VERSION : 0.1
   STRUCT
      CarrierNumber : Word;
      CarrierPosition : DWord;
      ActualSpeed : Word;
      CarrierDriveFaults : Word;
      CarrierDriveAlarms : Word;
      CarrierFaults : Word;
      Spare_Word : Word;
      RunningFWD : Bool;
      RunningREV : Bool;
      Stopped : Bool;
      ProductionHoldPB_Status : Bool;
      CrashDetectStatus : Bool;
      HeartBeat : Bool;
      AutoMode : Bool;
      ManualMode : Bool;
      IR_Remote_9_Pressed : Bool;
      EncoderCommFault : Bool;
      DriveCommFault : Bool;
      HMICommFault : Bool;
   END_STRUCT;
END_TYPE

TYPE "UDT_SDC_OUT"
VERSION : 0.1
   STRUCT
      Zone : Int;
      CarrierNum : Word;
      CarrierPosition : DWord;
      NextCarrierNum : Word;
      NextStopPos : DWord;
      DriveFwdCMD : Bool;
      DriveCmdSpeed : Word;
      Spare_Word_1 : Word;
      Spare_Word_2 : Word;
      HeartBeat : Bool;
      FaultReset : Bool;
      HighSpeedEnable : Bool;
      AtCmdPos : Bool;
      DuplicateCarrierNum : Word;
      FirstDuplicateFndPos : Bool;
      SecondDuplicateFndPos : Bool;
      Faults : "UDT_SDCOutFaults";
   END_STRUCT;
END_TYPE

TYPE "UDT_CarrierFaults"
VERSION : 0.1
   STRUCT
      Fault : Array[0..9] of Int;
   END_STRUCT;
END_TYPE

TYPE "UDT_SDC"
   STRUCT
      HMI : "UDT_Drive_HMI";
   END_STRUCT;
END_TYPE

TYPE "UDT_TrafficCop"
VERSION : 0.1
   STRUCT
      Element_1 : Bool;
      AutoSpeedFast : Word;
      AutoSpeedSlow : Word;
      CommandPosLowLimit : DWord;
      CommandPosHighLimit : DWord;
      CommandPos : DWord;
      AtCommandPos : Bool;
      DecelPosition : DWord;
   END_STRUCT;
END_TYPE

TYPE "UDT_SDC_6EMS_TS_STAT"
VERSION : 0.1
   STRUCT
      EMS : Array[1..6] of "UDT_SDC_EMS_TS_STAT";
   END_STRUCT;
END_TYPE

TYPE "UDT_SDC_6EMS_TS_STAT_HMI"
VERSION : 0.1
   STRUCT
      EMS : Array[1..6] of "UDT_SDC_EMS_TS_STAT_HMI";
   END_STRUCT;
END_TYPE

TYPE "UDT_EMS_IF_Q_VFC"
VERSION : 0.1
   STRUCT
      VFC_No : Byte;   // FU Nummer (z.B.: 1=Fahren, 2=Heben, 3=Schwenken) / VFC number (f.e.: 1=Drive, 2=Hoist, 3=Tilt)
      PW1 : Word;   // Prozesswort 1 / Processdataword 1
      PW2 : Word;   // Prozesswort 2 / Processdataword 2
      PW3 : Word;   // Prozesswort 3 / Processdataword 3
   END_STRUCT;
END_TYPE

TYPE "UDT_EMS_TA"
VERSION : 0.1
   STRUCT
      ZSW1 : Word;   // G120D Zustandswort 1 / Statusword 1
      ERROR : Word;   // G120D Störcode / Errorcode
      CURRENT : Word;   // G120D Strom / Current
      FAULT : Word;   // G120D Störcode / Errorcode
      ALARM : Word;
   END_STRUCT;
END_TYPE

TYPE "UDT_EMS_IF_Q_IQ"
VERSION : 0.1
   STRUCT
      BS1PH1_KANAL_1 : Bool;
      BS1PH1_KANAL_2 : Bool;
      BS1PH1_KANAL_3 : Bool;
      BS1PH1_KANAL_4 : Bool;
      BS1PH1_KANAL_5 : Bool;
      BS1PH1_KANAL_6 : Bool;
      BS1PH1_KANAL_7 : Bool;
      BS1PH1_KANAL_8 : Bool;
      BS1FC302 : Bool;
      AB1FCM1 : Bool;
      AB1QA1_R : Bool;
      I_1_3 : Bool;
      I_1_8 : Bool;
      I_1_5 : Bool;
      I_1_6 : Bool;
      I_1_7 : Bool;
      HE1BGS03a : Bool;
      HE1BGS03b : Bool;
      HE1BGS05 : Bool;
      BS1SFWE2 : Bool;
      I_2_4 : Bool;
      I_2_5 : Bool;
      I_2_6 : Bool;
      I_2_7 : Bool;
      I_6_0 : Bool;
      I_6_1 : Bool;
      I_6_2 : Bool;
      I_6_3 : Bool;
      I_6_4 : Bool;
      I_6_5 : Bool;
      I_6_6 : Bool;
      I_6_7 : Bool;
      "BS1PH1_L+" : Bool;
      BS1PH1_DAT : Bool;
      AB1QA1 : Bool;
      O_0_3 : Bool;
      O_0_4 : Bool;
      O_0_5 : Bool;
      O_0_6 : Bool;
      O_0_7 : Bool;
      HE1KK1 : Bool;
      O_8_1 : Bool;
      O_8_2 : Bool;
      O_8_3 : Bool;
      O_8_4 : Bool;
      O_8_5 : Bool;
      O_8_6 : Bool;
      O_8_7 : Bool;
      I_261_0 : Bool;
      I_261_1 : Bool;
      I_261_2 : Bool;
      I_261_3 : Bool;
      I_261_4 : Bool;
      I_261_5 : Bool;
      I_261_6 : Bool;
      I_261_7 : Bool;
      HE1BGG1 : Bool;
      "HE1BGG1:13" : Bool;
      HE1BGE05 : Bool;
      I_271_3 : Bool;
      I_271_4 : Bool;
      I_271_5 : Bool;
      I_271_6 : Bool;
      I_271_7 : Bool;
      SN1BGE04 : Bool;
      I_281_1 : Bool;
      I_281_2 : Bool;
      I_281_3 : Bool;
      I_281_4 : Bool;
      I_281_5 : Bool;
      I_281_6 : Bool;
      I_281_7 : Bool;
      I_285_0 : Bool;
      I_285_1 : Bool;
      I_285_2 : Bool;
      I_285_3 : Bool;
      I_285_4 : Bool;
      I_285_5 : Bool;
      I_285_6 : Bool;
      I_285_7 : Bool;
   END_STRUCT;
END_TYPE

TYPE "UDT_SDC_EMS_TS_STAT_HMI"
VERSION : 0.1
   STRUCT
      EMS_ID : Int;
      PROFILE : Int;
      DRIVE_POS : DInt;
      HOIST_POS : Int;
      ERROR : Int;
      "DRIVE_POS_%" : Int;
      SEK_NR : Int;
      STAT_1 : DWord;
      STAT_2 : Word;
      SORTE : DWord;
      FKT : DWord;
   END_STRUCT;
END_TYPE

TYPE "UDT_SDC_FT_STAT"
VERSION : 0.1
   STRUCT
      STAT : Array[1..4] of "UDT_SDC_EMS_TS_STAT";
   END_STRUCT;
END_TYPE

TYPE "UDT_EMS_IF_I"
VERSION : 0.1
   STRUCT
      EMS_ID : Int;   // EMS Nummer / EMS number
      CONT : "UDT_EMS_IF_I_CONTR";   // Steuerbit`s / Controlbit`s
      D_SETPOS : DInt;   // Sollposition Fahrantrieb / setpoint drive position (mm)
      D_SETSPEED : DInt;   // Sollgeschwindigkeit Fahrantrieb / set value drive speed (mm/min)
      H_SETPOS : Int;   // Sollposition Hubantrieb / setpoint hoist position (mm)
      H_SETSPEED : Int;   // Sollgeschwindigkeit Hubantrieb / setpoint hoist speed (mm/min)
      Reserve18 : Int;
      Reserve20 : Int;
      FB_VFC_No : Byte;   // Rückmeldung Prozesswerte FU`s / Feedback VFC PDAT
      FB_ER_WORD_No : Int;   // Rückmeldung Zähler Störnummern / Feedback Transfer counter error words
      DB_No : Int;   // DB Nummer Datentransfer / DB No. data transfer
      DBB_No : Int;   // DBB Nummer Datentransfer / DBB No. data transfer
      DB_UserData : DWord;   // Nutzdaten Datentransfer / User data, data transfer
      ERRORS_SPLC : "UDT_EMS_IF_I_SDC_ERRORS";   // Störungen Kopfsteuerung / Errors from System-PLC
      Reserve36 : Word;   // Reserve / spare
      Reserve38 : Word;   // Reserve / spare
   END_STRUCT;
END_TYPE

TYPE "UDT_EMS_PAR"
VERSION : 0.1
   STRUCT
      DRIVE : Struct
         Funct : Struct   // several functions
            Res0 : Bool := TRUE;   // Reserve: without swich-off Scanner
            IgnoreBridgeStopp : Bool := TRUE;   // Ignore Bridge Stopp-Position after Startpoint for Positioning
            DontIgnoreAPOSwhenDriving : Bool := FALSE;   // spare
            Speed0_1mm_s : Bool := FALSE;   // spare
            IR_noEMSnumber : Bool := FALSE;   // spare
            IR_noLogin : Bool := FALSE;   // spare
            Res6 : Bool := FALSE;   // spare
            Res7 : Bool := FALSE;   // spare
            Res8 : Bool := FALSE;   // spare
            Res9 : Bool := FALSE;   // spare
            Res10 : Bool := FALSE;   // spare
            Res11 : Bool := FALSE;   // spare
            Res12 : Bool := FALSE;   // spare
            Res13 : Bool := FALSE;   // spare
            Res14 : Bool := FALSE;   // spare
            Res15 : Bool := FALSE;   // spare
         END_STRUCT;
         V_FACT_1 : Real := 0.00266;
         V_SETP_1 : DInt := 600;   // Setpoint for calculation of factor
         V_FACT_2 : Real := 0.00246;
         V_SETP_2 : DInt := 3000;   // Setpoint for calculation of factor
         V_FACT_3 : Real := 0.00246;
         V_SETP_3 : DInt := 10000;   // Setpoint for calculation of factor
         V_FACT_4 : Real := 0.00236;
         V_SETP_4 : DInt := 20000;   // Setpoint for calculation of factor
         V_LIMIT_FACT : Real := 0.3;
         V_FACT_5 : Real := 0.00226;
         "V_FACT_ACT_V_<600" : Real := 0.0027;   // Factor for conversion of mm/min to U/min -> determined
         "V_FACT_ACT_V_<1200" : Real := 0.0027;   // Factor for conversion of mm/min to U/min -> determined
         V_min : DInt := 500;   // minimum speed in mm/min
         V_max_top : DInt := 36000;   // maximum speed if hoist raised in mm/min
         V_max_Not_top : DInt := 16000;   // maximum speed if hoist not raised in mm/min
         V_Pos_1_Reserve : DInt := 0;   // Positioning speed 1 / Positioning with position setpoint
         V_Pos_2 : DInt := 10000;   // Positioning speed 2 / Positioning with position setpoint
         V_Pos_3_Reserve : DInt := 12000;   // Positioning speed 3 / Positioning with position setpoint
         V_Fixed_1 : DInt := 3000;   // Fixed speed 1 in mm/min (IR manual)
         V_Fixed_2 : DInt := 13000;   // Fixed speed 2 in mm/min (IR manual)
         V_Fixed_3_Reserve : DInt := 18000;   // Fixed speed 3 in mm/min
         V_Fixed_4_SLS_SPEED : DInt := 15000;   // Fixed speed 4 in mm/min V_SafeSpeed
         V_DIV_FAST : DInt := 18000;   // speed for Divisor positioning fast
         DIV_POS_FAST : DInt := 40;   // Divisor to calculate braking distance for positioning fast (>=18m/min)
         DIV_POS_SLOW : DInt := 60;   // Divisor to calculate braking distance for positioning slow (<18m/min)
         TOL_SET_POS : Int := 2;   // tolerance (mm) for setting the position signal
         TOL_RESET_POS : Int := 6;   // tolerance (mm) for resetting the position signal
         Window_Pos : Int := 2;   // Window (mm) for shut-down during positioning
         Window_Overrun : Int := 6;   // Window (mm) for check "Stop Position overrun"
         Window_Pos_2 : Int := 800;   // Window (mm) for switching to positioning speed 2
         Window_Movement : Int := 10;   // Window (mm) for check "Movement without release"
         Window_Distance_Reserve : Int := 10;   // Window (mm) for distance controller
         Delay_Pos : Int := 2000;   // Delay EMS in position (ms)
         Reserve_118 : S5Time := S5T#5M;   // Delay Barcode scanner off
         Reserve_120 : S5Time := S5T#2M;   // Delay Barcode scanner on
         DelaySpeedContr : S5Time := S5T#9S_900MS;   // Delay for speed control
         TolSpeedContr : Int := 60;   // tolerance for speed control (in %)
         SYNCH_MID_VALUE : Int := 60;   // spare
         SYNCH_tINCREASE : Int := 30;
      END_STRUCT;
      Reserve : Array[1..5] of Word;
      HOIST : Struct
         V_Min : Int := 200;   // minimum speed in mm/min
         V_Max : Int := 8000;   // maximum speed in mm/min
         V_MaxOccLift : Int := 6600;   // maximum speed in mm/min occupied lifitng
         V_Reserve_2 : Int := 0;   // hoist speed spare
         V_Pos_1 : Int := 800;   // Positioning speed1
         V_Pos_2 : Int := 2000;   // Positioning speed 2
         V_Fixed_1 : Int := 2000;   // Fixed speed 1 in mm/min (IR manual)
         V_Fixed_2 : Int := 4000;   // Fixed speed 2 in mm/min (IR manual)
         V_Fixed_3_START : Int := 200;   // Fixed speed 3 in mm/min
         V_Fixed_4_SLS_SPEED : Int := 2000;   // Fixed speed 4 in mm/min
         V_Fixed_5_Reserve : Int := 2000;   // slow safe speed (2000)
         V_Fixed_6_SlowSpeed : Int := 4000;   // Global Speed paramter for TS {"DB_SDC_COMMAND".Section[1].Commands.hoist_slow}
         V_FACT_Hz_UP : Real := 0.01246;   // Factor for conversion of current value from converter in % to mm/min
         V_FACT_Hz_DOWN : Real := 0.01246;   // Factor for conversion of current value from converter in % to mm/min
         H_Window_POS_V1 : Int := 20;   // Window (mm) for switching to positioning speed 1
         H_Window_POS_V2 : Int := 140;   // Window (mm) for switching to positioning speed 2
         H_TOL_SET_POS : Int := 2;   // tolerance (mm) for setting the position signal
         H_TOL_RESET_POS : Int := 8;   // tolerance (mm) for resetting the position signal
         H_MIN : Int := 4;   // minimum height
         H_MIN_without_bypass : Int := 126;   // minimum height without bypass switch (120)
         H_REF_OFFSET : Int := 9;   // Offset to hoist position reference prox.switch
         H_REF : Int := 2641;   // Height reference initiator Position
         H_FACT_ENC1 : Real := 1.0;   // Factor for conversion of encoder value in mm / encoder 1
         H_FACT_ENC2 : Real := 1.0;   // Factor for conversion of encoder value in mm / encoder 2
         H_FACT_SPEED : Real := 0.316;   // Factor for conversion of encoder value / encoder 1or2 in mm for speed
         H_ENC_MAX_DIFF : Int := 50;   // maximum difference between encoders
         H_Slow : Int := 660;   // slow height (500)
         H_tIN_POS : Int := 1000;   // Delay HOIST in position (ms)
         H_REF_HMI : Int := 2641;   // Height HMI reference
      END_STRUCT;
      Reserve1 : Array[1..6] of Word;
      TILT : Array[1..34] of Word;
      Reserve2 : Array[1..6] of Word;
   END_STRUCT;
   // Reserve1[6] := 16#0000;
   // Reserve1[5] := 16#0000;
   // Reserve1[4] := 16#0000;
   // Reserve1[3] := 16#0000;
   // Reserve1[2] := 16#0000;
   // Reserve1[1] := 16#0000;
   // Reserve[5] := 16#0000;
   // Reserve[4] := 16#0000;
   // Reserve[3] := 16#0000;
   // Reserve[2] := 16#0000;
   // Reserve[1] := 16#0000;
   // Reserve2[1] := 16#0000;
   // Reserve2[2] := 16#0000;
   // Reserve2[3] := 16#0000;
   // Reserve2[4] := 16#0000;
   // Reserve2[5] := 16#0000;
   // Reserve2[6] := 16#0000;
END_TYPE

TYPE "UDT_TrafficCopCarrierStructure"
VERSION : 0.1
   STRUCT
      MoveFwd : Bool;
      DriveCmdSpeed : Word;
      CommandPos : DWord;
      AtCmdPos : Bool;
      NextStopPos : DWord;
      NextCarrierNumber : Word;
      CarrierNumber : Word;
   END_STRUCT;
END_TYPE

TYPE "UDT_TrafficCopZoneStructure"
VERSION : 0.1
   STRUCT
      Carrier : Array[0..99] of "UDT_TrafficCopCarrierStructure";
   END_STRUCT;
END_TYPE

TYPE "UDT_SDC_FT_COM"
VERSION : 0.1
   STRUCT
      COM : Array[1..7] of "UDT_SDC_EMS_TS_COM";
   END_STRUCT;
END_TYPE

TYPE "UDT_TC_ZoneMotion"
VERSION : 0.1
   STRUCT
      Zone : Array[0..60] of "UDT_ZnPosMotion";
   END_STRUCT;
END_TYPE

TYPE "UDT_TC_ZnPosMotion"
VERSION : 0.1
   STRUCT
      zone : Array[0..60] of "UDT_TrafficCopZnPosStructure";
   END_STRUCT;
END_TYPE

TYPE "UDT_ZnPosMotion"
VERSION : 0.1
   STRUCT
      ZonePos : Array[0..99] of "UDT_TrafficCopCarrierStructure";
   END_STRUCT;
END_TYPE

TYPE "UDT_HMIZonePositions"
   STRUCT
      ZonePosition : Word;
   END_STRUCT;
END_TYPE

TYPE "UDT_TC_SDCOutZone"
VERSION : 0.1
   STRUCT
      Carrier : Array[0..99] of "UDT_TC_SDCOutCarrier";
   END_STRUCT;
END_TYPE

TYPE "UDT_Drive_HMI"
   STRUCT
      G120D_STATUS : Word;
      G120D_CONTROL : Word;
   END_STRUCT;
END_TYPE

TYPE "UDT_TC_SDC_Out"
VERSION : 0.1
   STRUCT
      Zone : Array[0..60] of "UDT_TC_SDCOutZone";
   END_STRUCT;
END_TYPE

TYPE "UDT_TC_SDCOutCarrier"
VERSION : 0.1
   STRUCT
      DriveFwdCMD : Bool;
      DriveCmdSpeed : Int;
      NextStopPos : DWord;
      NextCarrierNum : Word;
      AtCmdPos : Bool;
   END_STRUCT;
END_TYPE

TYPE "UDT_IN"
   STRUCT
      G120D_CONTROL : "UDT_G120D_ZSW1_STATUS";
      G120D_STATUS : "UDT_G120D_STW1_CONTROL";
      DecrementCarrierIndex : Bool;
      IncrementCarrierIndex : Bool;
      CarrierStatusIndex : Int;
      DecrementStatusIndex : Bool;
      IncrementStatusIndex : Bool;
      DriveStatusIndex : Int;
      DecrementZoneIndex : Bool;
      IncrementZoneIndex : Bool;
      ZoneStatusIndex : Int;
   END_STRUCT;
END_TYPE

TYPE "UDT_TrafficCopZnPosStructure"
VERSION : 0.1
   STRUCT
      ZonePos : Array[0..40] of "UDT_TrafficCopZoneStructure";
   END_STRUCT;
END_TYPE

TYPE "UDT_ZoneStructure"
VERSION : 0.1
   STRUCT
      SpeedZoneStart : DWord;
      SpeedZoneEnd : DWord;
      Zone : Word;
      Description : String[10];
      Area : String[2];
      LastZone : Bool;
      StartPos : DWord;
      SpeedZone : Bool;
      NextZone : Int;
      PrevZone : Int;
      EndPos : DWord;
      AccumZone : Bool;
      ProductionZone : Bool;
      ProductionZoneSpacing : Word;
      MaxCarriers : Word;
      CarrierSpacing : Word;
      ClearToEnter : Bool;
      ClearOfStop : Bool;
      ClearZoneStart : Bool;
      ZoneFull : Bool;
      CarrierZnStatus : Array[0..60] of "UDT_ZoneCarrierStatus";
      CarrierZnStatusUnsorted : Array[0..60] of "UDT_ZoneCarrierStatus";
      InPositionTolerance : Word;
      NextCarrierClrHighSpeed : Word;
      DecelPositionOffset : Word;
      GapSpacingFault : Bool;
      GapFaultZnPosition : Int;
      GapFaultInZone : Int;
      FirstCarrierNumGapFlt : Int;
      SecondCarrierNumGapFlt : Int;
      FinePosStopZone : Bool;
      FineInPosTolerance : Word;
      FinePositionDecelOffset : Word;
      CoarseInPosTolerance : Word;
      CoarsePositionDecelOffset : Word;
      ZoneLength : Word;
      HMIZonePositionStatus : Array[1..20] of "UDT_HMIZonePositionStructure";
      HMIZonePositions : Array[1..20] of "UDT_HMIZonePositions";
      CarrierAtStop : Bool;
      CarrierNumAtStop : Word;
      StopControlFromEMS01 : "UDT_StopControlFromEMS01";
      ClearOfStopPos : DWord;
      StopStatusToEMS01 : "UDT_StopStatusToEMS01";
   END_STRUCT;
END_TYPE

TYPE "UDT_CarrierStructure"
VERSION : 0.1
   STRUCT
      SDC_IN : "UDT_SDC_IN";
      SDC_OUT : "UDT_SDC_OUT";
      ZoneFound : Word;
      Position : DWord;
      SpeedSelect : Word;
      MoveFWD : Bool;
      InProductionHold : Bool;
      Zone : Word;
      Area : String[2];
      AreaInt : Int;
      AutoSpeedFast : Word;
      AutoSpeedSlow : Word;
      InPositionTolerance : Word;
      DecelSpeed : Word;
      DecelStartPos : DWord;
      ZonePosition : Word;
      CommFlt : Bool;
      CarrierPosition : DWord;
      CarrierNumber : Word;
      FaultsMasked : Bool;
      Faulted : Bool;
   END_STRUCT;
END_TYPE

TYPE "UDT_Zone"
VERSION : 0.1
   STRUCT
      ZONE : Array[1..60] of "UDT_ZoneStructure";
   END_STRUCT;
END_TYPE

TYPE "UDT_ZoneCarrierStatus"
VERSION : 0.1
   STRUCT
      CarrierNumber : Word;
      Position : DWord;
      RunningFWD : Bool;
   END_STRUCT;
END_TYPE

TYPE "UDT_OUT"
   STRUCT
      DecrementCarrierIndex : Bool;
      IncrementCarrierIndex : Bool;
      CarrierStatusIndex : Int;
      DecrementStatusIndex : Bool;
      IncrementStatusIndex : Bool;
      DriveStatusIndex : Int;
      DecrementZoneIndex : Bool;
      IncrementZoneIndex : Bool;
      ZoneStatusIndex : Int;
   END_STRUCT;
END_TYPE

TYPE "UDT_Carrier_Drive_Data"
   STRUCT
      CARRIER : Array[1..99] of "UDT_Drive_Data";
   END_STRUCT;
END_TYPE

TYPE "UDT_Drive_Data"
   STRUCT
      Drive_Control : Word;
      Drive_Status : Word;
   END_STRUCT;
END_TYPE

TYPE "UDT_Carrier_IO_HMI"
   STRUCT
      Carrier_Slot02_Inputs : Byte;
      Carrier_Slot03_Outputs : Byte;
      Carrier_Slot04_Inputs : Word;
      Carrier_Slot05_Outputs : Word;
   END_STRUCT;
END_TYPE

TYPE "UDT_IO_Data"
   STRUCT
      Slot2SafeInputs : Byte;
      Slot3SafeOutputs : Byte;
      Slot4StdInputs : Word;
      Slot5StdOutputs : Word;
   END_STRUCT;
END_TYPE

TYPE "UDT_Carrier_IO_Data"
   STRUCT
      CARRIER : Array[1..99] of "UDT_IO_Data";
   END_STRUCT;
END_TYPE

TYPE "UDT_Carrier_Status_HMI"
   STRUCT
      CarrierPosition : DWord;
      ActualSpeed : Word;
      RunningFWD : Bool;
      RunningREV : Bool;
      ProductionHoldPB_Status : Bool;
      CrashDetectStatus : Bool;
      AutoMode : Bool;
      ManualMode : Bool;
      DriveFwdCMD : Bool;
      DriveCmdSpeed : Word;
      NextCarrierNum : Word;
      NextStopPosition : DWord;
      Zone : Int;
      Area : String[2];
      CarrierFaultCode : Int;
      AtCmdPos : Bool;
      CommFlt : Bool;
      Faulted : Bool;
      CarrierStatusIndex : Int;
      DriveStatusIndex : Int;
      ZoneStatusIndex : Int;
      EncoderCommFault : Bool;
      DriveCommFault : Bool;
      HMICommFault : Bool;
      SetMaskCarrierFaultsPB : Bool;
      MaskCarrierFaultsLT : Bool;
      ResetMaskCarrierFaultsPB : Bool;
   END_STRUCT;
END_TYPE

TYPE "UDT_Zone_Status_HMI"
   STRUCT
      ZoneIndex : Int;
      ZoneType : String;
      PrevZoneNumber : Int;
      NextZoneNumber : Int;
      ZoneStartPosition : DWord;
      ZoneEndPosition : DWord;
      ZoneFull : Bool;
      AccumZone : Bool;
      ProdZone : Bool;
      SpeedZone : Bool;
      SpeedZoneStartPos : DWord;
      SpeedZoneEndPos : DWord;
      AccumZoneSpacing : Word;
      ProductionZoneSpacing : Word;
      CarrierZoneStatus : Array[0..60] of "UDT_ZoneCarrierStatus";
   END_STRUCT;
END_TYPE

TYPE "UDT_StopStatusToEMS01"
VERSION : 0.1
   STRUCT
      CarrierInStop : Bool;
      Blocked : Bool;
      CarrierBlockZoneClear : Bool;
      CycleComplete : Bool;
      CarrierPositComp : Bool;
      CarrierMoving : Bool;
      CarrierAutoInStop : Bool;
      Spare_11 : Bool;
      Spare_12 : Bool;
      Spare_13 : Bool;
      Spare_14 : Bool;
      StopFaultReady : Bool;
   END_STRUCT;
END_TYPE

TYPE "UDT_StopControlFromEMS01"
VERSION : 0.1
   STRUCT
      HoldStop : Bool;
      SetToRelease : Bool;
      DrivePermit : Bool;
      BypassStop : Bool;
      PowerX_FER_Set_ToExit : Bool;
      SpareBool3 : Bool;
      SpareBool4 : Bool;
      SpareBool5 : Bool;
      SpareBool6 : Bool;
      SpareBool7 : Bool;
      SpareBool8 : Bool;
      SpareBool9 : Bool;
      SpareBool10 : Bool;
      SpareBool11 : Bool;
      SpareBool12 : Bool;
      SpareBool13 : Bool;
      SpareBool14 : Bool;
      SpareBool15 : Bool;
   END_STRUCT;
END_TYPE

TYPE "UDT_G120D_STW1_CONTROL"
VERSION : 0.1
   STRUCT
      Bit_08_JOG_R : Bool;   // 1=tippen rechtsseitig EIN/ 0= AUS / 1=jogging on right-hand side ON/ 0= OFF
      Bit_09_JOG_L : Bool;   // 1=tippen linksseitig EIN/ 0= AUS / 1=jogging on left-hand side ON/ 0= OFF
      Bit_10_CONTR_PLC : Bool;   // 1=Bedienung über PLC erforderlich/ 0=keine Bedienung über PLC erforderlich / 1=control by PLC required/ 0=no control by PLC required
      Bit_11_REVERSE : Bool;   // 1=Umkehrung des Sollwerts/ 0=keine Umkehrung / 1=inversion of setpoint/ 0=no inversion of setpoint
      Bit_12_BRAKE_Release : Bool;   // 1= Löse Bremse / 1= Release Break / 1= Manual Brake Release
      Bit_13_DDS : Bool;   // 1=DDS1 FU Datenset / 0=DDS0 FU Datenset / 1=DDS1 FU Dataset / 0=DDS0 FU Dataset
      Bit_14_DO0 : Bool;   // 1=Digitaler Ausgang aktiv/ 0=Digitaler Ausgang nicht aktiv / 1=Digital Output activ/ 0=Digital Output not activ
      Bit_15_DO1 : Bool;   // 1=Digitaler Ausgang aktiv/ 0=Digitaler Ausgang nicht aktiv / 1=Digital Output activ/ 0=Digital Output not activ
      Bit_00_ON : Bool;   // 1=EIN/ 0=AUS / 1=ON/ 0=OFF2
      Bit_01_AUS2_INH : Bool;   // 1=Betriebsvoraussetzung/ 0=AUS2 - Pulsverzögerer, Spannung auf einmal aus / 1=operation condition/ 0=AUS2 - pulse inhibitor, voltage off at once
      Bit_02_AUS3_STOP : Bool;   // 1=Betriebsvoraussetzung / 0=AUS3 - schneller Halt / 1=operation condition / 0=AUS3 - fast stop
      Bit_03_EN : Bool;   // 1=Freigabe Betrieb/ 0=deaktiviere Betrieb / 1=enable operation/ 0=disable operation
      Bit_04_EN_RAMP : Bool;   // 1=1=Betriebsvoraussetzung / 0=deaktiviere Funktionsrampengenerator / 1=operation condition / 0=disable ramp function generator
      Bit_05_START_RAMP : Bool;   // 1=Aktiviere Rampenfunktion / 0=deaktivere RFG / 1=enable ramp function generator / 0=stoppen RFG
      Bit_06_SETPOINT : Bool;   // 1=Freigabe Sollwert/ 0=deaktiviere Sollwert / 1=enable setpoint/ 0=disable setpoint
      Bit_07_RESET : Bool;   // 1=Störung quittieren / 0= irrelevant / 1=Reset fault / 0= irrelevant
   END_STRUCT;
END_TYPE

TYPE "UDT_G120D_ZSW1_STATUS"
VERSION : 0.1
   STRUCT
      Bit_08_NO_DEVIATION : Bool;   // 1=keine Abweichung des Sollwerts / 0=Abweichung / 1=no deviation current-setpoint / 0=deviation / Setpoint / actual value deviation within the tolerance range.
      Bit_09_CONTR_PLC : Bool;   // 1=Kontrolle über PLC erforderlich/ 0=keine Kontrolle erforderlich / 1=control by PLC required/ 0=no control by PLC required / The automation system is requested to ac-cept the inverter control.
      Bit_10_F_MAX : Bool;   // 1=fmax erreicht/ 0= unter fmax / 1=fmax reached/ 0= below fmax / Speed is greater than or equal to the corre-sponding maximum speed.
      Bit_11_LIMIT_REACHED : Bool;   // 1=keine Warnung/ 0=Warnung: Motor an Spannungsgrenze / 1=no warning/ 0=warning:Motor at limit of current / Comparison value for current or torque has been reached or exceeded.
      Bit_12_BRAKE_OPEN : Bool;   // 1= / 0=Haltebremse / motor Brake is open
      Bit_13_NO_OVERTEMP : Bool;   // 1= / 0=Motorüberlast / Drive Overtemperature
      Bit_14_CW_CCW : Bool;   // 1=Rechtslauf/ 0=Linkslauf / On for drive runnin clockwise/off counterclockwise
      Bit_15_OVERL : Bool;   // 1= /0= Konvertierer Überlast / 1= /0= Konverter overload / 0 = Alarm, in-verter thermal overload/on CDS display
      Bit_00_READY_RUN : Bool;   // 1=bereit zum betreiben/ 0= nicht bereit / 1=ready to run/ 0= not ready to run / Power supply switched on; electronics initial-ized; pulses locked.
      Bit_01_READY_ON : Bool;   // 1=bereit zum einschalten/ 0= nicht bereit / 1=ready to switch on/ 0= not ready to switch on / Motor is switched on (ON/OFF1 = 1), no fault is active. With the command "Enable opera-tion" (STW1.3), the inverter switches on the motor.
      Bit_02_ENABLE : Bool;   // 1=Freigabe Bedienung / 0=deaktiviere Bedienung / 1=operation enabled / 0=operation disabled / Motor follows setpoint. See control word 1, bit 3.
      Bit_03_FAULT : Bool;   // 1=Störung / 0=keine Störung / 1=fault / 0=no fault / The inverter has a fault. Acknowledge fault using STW1.7
      Bit_04_OFF2 : Bool;   // 1=kein AUS2 / 0=AUS2 Befehl ist vorhanden / 1=no AUS2 / 0=AUS2 command is present / OFF2 Coast down to standstill is not active.
      Bit_05_OFF3 : Bool;   // 1=kein AUS3 / 0=AUS3 Befehl ist vorhanden / 1=no AUS3 / 0=AUS3 command is present / OFF3 Quick stop is not active.
      Bit_06_LOCK_OUT : Bool;   // 1=sperre Ausschaltung / 0=keine Sperrung / 1=closing lock-out / 0=no closing lock-out / It is only possible to switch on the motor after an OFF1 followed by ON.
      Bit_07_WARN : Bool;   // 1=Warnung / 0= keine Warnung / 1=Warning / 0= no warning
   END_STRUCT;
END_TYPE

TYPE "UDT_G120D_ERRORS"
VERSION : 0.1
   STRUCT
      F_X33_F1 : Bool;   // Fehler Überstrom
      F_X34_F2 : Bool;   // Fehler Überspannung
      F_X35_F3 : Bool;   // Fehler Unterspannung
      F_X36_F4 : Bool;   // Fehler Inverter Übertemperatur
      F_X37_F41 : Bool;   // Fehler Motordatenerkennung
      F_X38_F52 : Bool;   // Fehler Leistungsteil
      F_X39_F62 : Bool;   // Fehler MMC Daten sind fehlerhaft
      F_X40_F70 : Bool;   // Fehler PLC Sollposition
      F_X41_F71 : Bool;   // Fehler USS Sollposition, Überwachung
      F_X42_F72 : Bool;   // Fehler USS Sollposition, USS Master
      F_X43_F90 : Bool;   // Fehler Gebersignal
      F_X44_F395 : Bool;   // Fehler CU/PM wechsel
      bit_14 : Bool;   // Reserve
      bit_15 : Bool;   // Reserve
      bit_16 : Bool;   // Reserve
      bit_17 : Bool;   // Reserve
   END_STRUCT;
END_TYPE

TYPE "UDT_SDC_EMS_FLAGS"
VERSION : 0.1
   STRUCT
      PRESENT : Bool;   // EMS vorhanden
      IN_HW : Bool;   // EMS in HardwareConfiguration
      ACTIV : Bool;   // EMS activiert
      ENABLE : Bool;   // EMS enable
      COMM_FAULT : Bool;   // EMS communicationsfehler
      FAULTY : Bool;   // EMS fehlerhaft
      SIMULATION : Bool;   // EMS simualtion
      Spare_0_7 : Bool;   // Spare
      Spare_1_0 : Bool;   // Spare
      Spare_1_1 : Bool;   // Spare
      Spare_1_2 : Bool;   // Spare
      Spare_1_3 : Bool;   // Spare
      Spare_1_4 : Bool;   // Spare
      Spare_1_5 : Bool;   // Spare
      Spare_1_6 : Bool;   // Spare
      Spare_1_7 : Bool;   // Spare
   END_STRUCT;
END_TYPE

TYPE "UDT_SDC_TS_PARAMETER"
VERSION : 0.1
   STRUCT
      ALLG : "UDT_SDC_TS_PAR_ALLG";   // allgemeine Sections Parameter
      PROFIL : Array[1..10] of "UDT_SDC_TS_PAR_PROFIL";   // Profilbezogene Sections Parameter
   END_STRUCT;
END_TYPE

TYPE "UDT_SDC_TS_PAR_PROFIL"
VERSION : 0.1
   STRUCT
      Hoist_Pos_start : Int;   // Start of hoist positioning; offset from start pos.(mm)
      Height : Int := 2651;   // Setpoint: hoist position (mm)
      Hoist_speed : Int := 2000;   // Setpoint: hoist speed (mm/min)
      Hoist_offset_1 : Int;   // set value: hoist offset (mm)
      Hoist_offset_2 : Int;   // set value: hoist offset (mm)
      Hoist_offset_3 : Int;   // set value: hoist offset (mm)
      Hoist_offset_4 : Int;   // set value: hoist offset (mm)
      Hoist_Start_offset_1 : Int;   // Start der Hubbewegung zu offset 1, Offset von Startpos. (mm)
      Hoist_Start_offset_2 : Int;   // Start der Hubbewegung zu offset 1, Offset von Startpos. (mm)
      Hoist_Start_offset_3 : Int;   // Start der Hubbewegung zu offset 1, Offset von Startpos. (mm)
      Hoist_Start_offset_4 : Int;   // Start der Hubbewegung zu offset 1, Offset von Startpos. (mm)
   END_STRUCT;
END_TYPE

TYPE "UDT_SDC_TS_PAR_ALLG"
VERSION : 0.1
   STRUCT
      SEK_NEXT_1 : Int;   // Sektion next 1
      SEK_NEXT_2 : Int;   // Sektion next 2
      Spare : Array[4..5] of Byte;   // Spare
      POS : "UDT_SDC_TS_PAR_POS";   // Pos Parameter
      FLAGS : Struct
         DIST_VAL : Array[0..15] of Bool;   // Abstandswerte
         one_profile : Bool;   // Reserved for: only one profile
         BLIND : Bool;   // Reserved for: Blind travel without position values
         NO_DIST_CONT : Bool;   // without distance control (no slow speed, ...)
         SYNCH_AREA : Bool;   // synchronous conveyor area
         bit24 : Bool;   // spare
         bit25 : Bool;   // spare
         bit26 : Bool;   // spare
         bit27 : Bool;   // spare
         EN_HOIST : Bool;   // Hoist/tilt enable
         D_RESET_AFTER : Bool;   // Antrieb belegt nach Reset vorhanden
         D_PULK : Bool;   // Antriebs PULK
         bit33 : Bool;   // spare
         bit34 : Bool;   // spare
         bit35 : Bool;   // spare
         bit36 : Bool;   // spare
         Deutronic_ON : Bool;   // Reserved for: DEUTRONIC CHARGE COMPUTER ON
      END_STRUCT;
      Stop_Position : Int;   // Stopp position, offset from start pos.(mm)
      Drive_speed_1 : DInt;   // set value: drive speed (mm/min)
      Drive_speed_2 : DInt;   // set value: drive speed (mm/min)
   END_STRUCT;
   // FLAGS.DIST_VAL[0] := true;
END_TYPE

TYPE "UDT_SDC_TS_PAR_POS"
VERSION : 0.1
   STRUCT
      Start_1 : DInt := 0;   // mm
      End_1 : DInt := 0;   // mm
      Start_2 : DInt;   // Reserve
      End_2 : DInt;   // Reserve
      Actionpoint_1 : Int;   // Fahrantrieb Aktionspunkt 1
      Actionpoint_2 : Int;   // Fahrantrieb Aktionspunkt 2
   END_STRUCT;
END_TYPE

TYPE "UDT_EMS_IF_Q"
VERSION : 0.1
   STRUCT
      STAT : "UDT_EMS_IF_Q_STAT";   // Statusbit`s / Stausbit`s
      ERROR : Int;   // Störnummer / Error number
      D_POS : DInt;   // Fahrantrieb Position in mm / Drive position in mm
      H_POS : Int;   // Hubantrieb Position in mm / Hoist position in mm
      SPARE_POS : Int;
      VFC : "UDT_EMS_IF_Q_VFC";   // Prozesswerte FU`s / Processdata VFC
      IQ : "UDT_EMS_IF_Q_IQ";   // Ein-Ausgänge / In-Outputs
      ER_WORD_No : Int;   // Zähler Störnummern / Counter error words
      ER_WORD : Word;   // Datenwort Störnummern / Dataword error words
      FB_DBNo : Int;   // Rückmeldung DB Nummer Datentransfer / Feedback DB No. data transfer
      FB_DBBNo : Int;   // Rückmeldung DBB Nummer Datentransfer / Feedback DBB No. data transfer
   END_STRUCT;
END_TYPE

TYPE "UDT_SDC_EMS"
VERSION : 0.1
   STRUCT
      IF_I_EMS : "UDT_EMS_IF_Q";   // Inputs from EMS
      IF_Q_EMS : "UDT_EMS_IF_I";   // Outputs to EMS
      TS_PAR : Struct   // Section parameters
         ALLG : "UDT_SDC_TS_PAR_ALLG";   // Section parameters allg
         PROFIL : "UDT_SDC_TS_PAR_PROFIL";   // Section parameters Profil
      END_STRUCT;
      TS_STAT : "UDT_SDC_EMS_TS_STAT";   // EMS Sektion Stat Daten
      TS_COM : "UDT_SDC_EMS_TS_COM";   // EMS Sektion Com Daten
      FKT : "UDT_SDC_EMS_FKT_BITs";   // EMS Funktionen
      FKT_RESET : "UDT_SDC_EMS_FKT_BITs";   // EMS Funktionen reset
      FLAGS : "UDT_SDC_EMS_FLAGS";   // EMS Fahnen
      FKT_INFO_REP_1 : Int;   // EMS Funktionen Info Repair 1
      FKT_INFO_REP_2 : Int;   // EMS Funktionen Info Repair 2
      PROFIL : Int;   // Profile Number
      CYCLE_COUNTER : Int;   // Zykluszähler
      PRECEDING_EMS : Int;   // preciding EMS
      DISTANCE : DInt;   // Abstand zum vorangehenden EMS
      ABS_POS : DInt;   // absolute Positon
      NewSektion : Bool;   // New Sektion
      BcOk : Bool;   // Barcode ist OK
      SekOk : Bool;   // Sektion is OK
      Spare_0_3 : Bool;   // Spare
      Spare_0_4 : Bool;   // Spare
      Spare_0_5 : Bool;   // Spare
      Spare_0_6 : Bool;   // Spare
      Spare_0_7 : Bool;   // Spare
      Send_EMS_PAR_Act : Bool;   // Sende EMS Parameter aktiv
      Send_EMS_PAR_End : Bool;   // Sende EMS Parameter ende
      Send_EMS_LEAPS_Act : Bool;   // Sende EMS Sprünge aktiv
      Send_EMS_LEAPS_End : Bool;   // Sende EMS Sprünge ende
      H_C_Pos : Array[0..4] of Bool;   // Hub Kommando positionierung / Offset 1 / ,...
      Spare246 : Array[246..249] of Byte;   // Spare
      ER : "UDT_EMS_IF_I_SDC_ERRORS";
      WA_DIST : Bool;   // Warning Distance
      WA_COLL : Bool;   // Warning Collision Sensor activ
      WA_DIST_SAFETY : Bool;   // Warning Distance safety
      WA_Spare_2_3 : Bool;   // Warning Spare 2.3
      WA_Spare_2_4 : Bool;   // Warning Spare 2.4
      WA_Spare_2_5 : Bool;   // Warning Spare 2.5
      WA_Spare_2_6 : Bool;   // Warning Spare 2.6
      WA_Spare_2_7 : Bool;   // Warning Spare 2.7
      WA_Spare_3 : Byte;   // Warning Spare 3
      Spare254 : Array[254..257] of Byte;   // Spare
      VersNo : Array[0..1] of Byte;
   END_STRUCT;
END_TYPE

TYPE "UDT_SDC_EMS_TS_STAT"
VERSION : 0.1
   STRUCT
      VAL : "UDT_SDC_TS_IF_STATUS_VAL";
      BIT : "UDT_SDC_TS_IF_STATUS_BIT";
      SORTE : Array[1..4] of Char;   // Karossentyp
      FKT : "UDT_SDC_EMS_FKT_BITs";
      SPARE : Word;
   END_STRUCT;
END_TYPE

